      ProcessValue <- "Perfiladores\Perfilador.PL1_1"
   IOField "Champ E/S_115" at 543,307 size 51x25; FormatPattern s999999
      Appearance <- "Perfiladores\Perfilador.PresenciaPieza"
      ProcessValue <- "Perfiladores\Perfilador.PL1_2"
   IOField "Champ E/S_116" at 543,328 size 51x24; FormatPattern s999999
      Appearance <- "Perfiladores\Perfilador.PresenciaPieza"
      ProcessValue <- "Perfiladores\Perfilador.PL2_1"
   IOField "Champ E/S_117" at 543,347 size 51x25; FormatPattern s999999
      Appearance <- "Perfiladores\Perfilador.PresenciaPieza"
      ProcessValue <- "Perfiladores\Perfilador.PL2_2"
   TextField "Campo de texto_123" at 503,310 size 35x18; Text 'PL1-2'
   TextField "Campo de texto_124" at 503,331 size 35x18; Text 'PL2-1'
   TextField "Campo de texto_125" at 503,350 size 35x18; Text 'PL2-2'
   TextField "Campo de texto_134" at 328,210 size 17x18; Text 'F1'
   IOField "Champ E/S_126" at 352,207 size 51x25; FormatPattern s999999
      Appearance <- "Rolos\Rolos.PresenciaPieza"
      ProcessValue <- "Rolos\Rolos.F1"
   IOField "Champ E/S_127" at 352,227 size 51x25; FormatPattern s999999
      Appearance <- "Rolos\Rolos.PresenciaPieza"
      ProcessValue <- "Rolos\Rolos.F2"
   IOField "Champ E/S_128" at 352,248 size 51x24; FormatPattern s999999
      Appearance <- "Rolos\Rolos.PresenciaPieza"
      ProcessValue <- "Rolos\Rolos.F3"
   IOField "Champ E/S_129" at 352,267 size 51x25; FormatPattern s999999
      Appearance <- "Rolos\Rolos.PresenciaPieza"
      ProcessValue <- "Rolos\Rolos.F4"
   TextField "Campo de texto_135" at 328,229 size 17x18; Text 'F2'
   TextField "Campo de texto_136" at 328,249 size 17x18; Text 'F3'
   TextField "Campo de texto_137" at 328,269 size 17x18; Text 'F4'
   TextField "Campo de texto_138" at 328,290 size 35x18; Text 'PL1-1'
   IOField "Champ E/S_130" at 368,287 size 51x25; FormatPattern s999999
      Appearance <- "Rolos\Rolos.PresenciaPieza"
      ProcessValue <- "Rolos\Rolos.PL1_1"
   IOField "Champ E/S_131" at 368,307 size 51x25; FormatPattern s999999
      Appearance <- "Rolos\Rolos.PresenciaPieza"
      ProcessValue <- "Rolos\Rolos.PL1_2"
   IOField "Champ E/S_132" at 368,328 size 51x24; FormatPattern s999999
      Appearance <- "Rolos\Rolos.PresenciaPieza"
      ProcessValue <- "Rolos\Rolos.PL2_1"
   IOField "Champ E/S_133" at 368,347 size 51x25; FormatPattern s999999
      Appearance <- "Rolos\Rolos.PresenciaPieza"
      ProcessValue <- "Rolos\Rolos.PL2_2"
   TextField "Campo de texto_139" at 328,310 size 35x18; Text 'PL1-2'
   TextField "Campo de texto_140" at 328,331 size 35x18; Text 'PL2-1'
   TextField "Campo de texto_141" at 328,350 size 35x18; Text 'PL2-2'
   TextField "Campo de texto_142" at 151,210 size 17x18; Text 'F1'
   IOField "Champ E/S_134" at 175,207 size 51x25; FormatPattern s999999
      Appearance <- "Araña\Araña.PresenciaPieza"
      ProcessValue <- "Araña\Araña.F1"
   IOField "Champ E/S_135" at 175,227 size 51x25; FormatPattern s999999
      Appearance <- "Araña\Araña.PresenciaPieza"
      ProcessValue <- "Araña\Araña.F2"
   IOField "Champ E/S_136" at 175,248 size 51x24; FormatPattern s999999
      Appearance <- "Araña\Araña.PresenciaPieza"
      ProcessValue <- "Araña\Araña.F3"
   IOField "Champ E/S_137" at 175,267 size 51x25; FormatPattern s999999
      Appearance <- "Araña\Araña.PresenciaPieza"
      ProcessValue <- "Araña\Araña.F4"
   TextField "Campo de texto_143" at 151,229 size 17x18; Text 'F2'
   TextField "Campo de texto_144" at 151,249 size 17x18; Text 'F3'
   TextField "Campo de texto_145" at 151,269 size 17x18; Text 'F4'
   TextField "Campo de texto_146" at 151,290 size 35x18; Text 'PL1-1'
   IOField "Champ E/S_138" at 191,287 size 51x25; FormatPattern s999999
      Appearance <- "Araña\Araña.PresenciaPieza"
      ProcessValue <- "Araña\Araña.PL1_1"
   IOField "Champ E/S_139" at 191,307 size 51x25; FormatPattern s999999
      Appearance <- "Araña\Araña.PresenciaPieza"
      ProcessValue <- "Araña\Araña.PL1_2"
   IOField "Champ E/S_140" at 191,328 size 51x24; FormatPattern s999999
      Appearance <- "Araña\Araña.PresenciaPieza"
      ProcessValue <- "Araña\Araña.PL2_1"
   IOField "Champ E/S_141" at 191,347 size 51x25; FormatPattern s999999
      Appearance <- "Araña\Araña.PresenciaPieza"
      ProcessValue <- "Araña\Araña.PL2_2"
   TextField "Campo de texto_147" at 151,310 size 35x18; Text 'PL1-2'
   TextField "Campo de texto_148" at 151,331 size 35x18; Text 'PL2-1'
   TextField "Campo de texto_149" at 151,350 size 35x18; Text 'PL2-2'
   TextField "Campo de texto_150" at 679,210 size 17x18; Text 'F1'
   IOField "Champ E/S_142" at 703,207 size 51x25; FormatPattern s999999
      Appearance <- "Cinta\Cinta.PresenciaPieza"
      ProcessValue <- "Cinta\Cinta.F1"
   IOField "Champ E/S_143" at 703,227 size 51x25; FormatPattern s999999
      Appearance <- "Cinta\Cinta.PresenciaPieza"
      ProcessValue <- "Cinta\Cinta.F2"
   IOField "Champ E/S_144" at 703,248 size 51x24; FormatPattern s999999
      Appearance <- "Cinta\Cinta.PresenciaPieza"
      ProcessValue <- "Cinta\Cinta.F3"
   IOField "Champ E/S_145" at 703,267 size 51x25; FormatPattern s999999
      Appearance <- "Cinta\Cinta.PresenciaPieza"
      ProcessValue <- "Cinta\Cinta.F4"
   TextField "Campo de texto_151" at 679,229 size 17x18; Text 'F2'
   TextField "Campo de texto_152" at 679,249 size 17x18; Text 'F3'
   TextField "Campo de texto_153" at 679,269 size 17x18; Text 'F4'
   TextField "Campo de texto_154" at 679,290 size 35x18; Text 'PL1-1'
   IOField "Champ E/S_146" at 719,287 size 51x25; FormatPattern s999999
      Appearance <- "Cinta\Cinta.PresenciaPieza"
      ProcessValue <- "Cinta\Cinta.PL1_1"
   IOField "Champ E/S_147" at 719,307 size 51x25; FormatPattern s999999
      Appearance <- "Cinta\Cinta.PresenciaPieza"
      ProcessValue <- "Cinta\Cinta.PL1_2"
   IOField "Champ E/S_148" at 719,328 size 51x24; FormatPattern s999999
      Appearance <- "Cinta\Cinta.PresenciaPieza"
      ProcessValue <- "Cinta\Cinta.PL2_1"
   IOField "Champ E/S_149" at 719,347 size 51x25; FormatPattern s999999
      Appearance <- "Cinta\Cinta.PresenciaPieza"
      ProcessValue <- "Cinta\Cinta.PL2_2"
   TextField "Campo de texto_155" at 679,310 size 35x18; Text 'PL1-2'
   TextField "Campo de texto_156" at 679,331 size 35x18; Text 'PL2-1'
   TextField "Campo de texto_157" at 679,350 size 35x18; Text 'PL2-2'
   TextField "Campo de texto_158" at 851,210 size 17x18; Text 'F1'
   IOField "Champ E/S_150" at 875,207 size 51x25; FormatPattern s999999
      Appearance <- "Pinza\Pinza.PresenciaPieza"
      ProcessValue <- "Pinza\Pinza.F1"
   IOField "Champ E/S_151" at 875,227 size 51x25; FormatPattern s999999
      Appearance <- "Pinza\Pinza.PresenciaPieza"
      ProcessValue <- "Pinza\Pinza.F2"
   IOField "Champ E/S_152" at 875,248 size 51x24; FormatPattern s999999
      Appearance <- "Pinza\Pinza.PresenciaPieza"
      ProcessValue <- "Pinza\Pinza.F3"
   IOField "Champ E/S_153" at 875,267 size 51x25; FormatPattern s999999
      Appearance <- "Pinza\Pinza.PresenciaPieza"
      ProcessValue <- "Pinza\Pinza.F4"
   TextField "Campo de texto_159" at 851,229 size 17x18; Text 'F2'
   TextField "Campo de texto_160" at 851,249 size 17x18; Text 'F3'
   TextField "Campo de texto_161" at 851,269 size 17x18; Text 'F4'
   TextField "Campo de texto_162" at 851,290 size 35x18; Text 'PL1-1'
   IOField "Champ E/S_154" at 891,287 size 51x25; FormatPattern s999999
      Appearance <- "Pinza\Pinza.PresenciaPieza"
      ProcessValue <- "Pinza\Pinza.PL1_1"
   IOField "Champ E/S_155" at 891,307 size 51x25; FormatPattern s999999
      Appearance <- "Pinza\Pinza.PresenciaPieza"
      ProcessValue <- "Pinza\Pinza.PL1_2"
   IOField "Champ E/S_156" at 891,328 size 51x24; FormatPattern s999999
      Appearance <- "Pinza\Pinza.PresenciaPieza"
      ProcessValue <- "Pinza\Pinza.PL2_1"
   IOField "Champ E/S_157" at 891,347 size 51x25; FormatPattern s999999
      Appearance <- "Pinza\Pinza.PresenciaPieza"
      ProcessValue <- "Pinza\Pinza.PL2_2"
   TextField "Campo de texto_163" at 851,310 size 35x18; Text 'PL1-2'
   TextField "Campo de texto_164" at 851,331 size 35x18; Text 'PL2-1'
   TextField "Campo de texto_165" at 851,350 size 35x18; Text 'PL2-2'
   TextField "Campo de texto_166" at 1029,210 size 17x18; Text 'F1'
   IOField "Champ E/S_158" at 1053,207 size 51x25; FormatPattern s999999
      Appearance <- "Plegadora\Plegadora.PresenciaPieza"
      ProcessValue <- "Plegadora\Plegadora.F1"
   IOField "Champ E/S_159" at 1053,227 size 51x25; FormatPattern s999999
      Appearance <- "Plegadora\Plegadora.PresenciaPieza"
      ProcessValue <- "Plegadora\Plegadora.F2"
   IOField "Champ E/S_160" at 1053,248 size 51x24; FormatPattern s999999
      Appearance <- "Plegadora\Plegadora.PresenciaPieza"
      ProcessValue <- "Plegadora\Plegadora.F3"
   IOField "Champ E/S_161" at 1053,267 size 51x25; FormatPattern s999999
      Appearance <- "Plegadora\Plegadora.PresenciaPieza"
      ProcessValue <- "Plegadora\Plegadora.F4"
   TextField "Campo de texto_167" at 1029,229 size 17x18; Text 'F2'
   TextField "Campo de texto_168" at 1029,249 size 17x18; Text 'F3'
   TextField "Campo de texto_169" at 1029,269 size 17x18; Text 'F4'
   TextField "Campo de texto_170" at 1029,290 size 35x18; Text 'PL1-1'
   IOField "Champ E/S_162" at 1069,287 size 51x25; FormatPattern s999999
      Appearance <- "Plegadora\Plegadora.PresenciaPieza"
      ProcessValue <- "Plegadora\Plegadora.PL1_1"
   IOField "Champ E/S_163" at 1069,307 size 51x25; FormatPattern s999999
      Appearance <- "Plegadora\Plegadora.PresenciaPieza"
      ProcessValue <- "Plegadora\Plegadora.PL1_2"
   IOField "Champ E/S_164" at 1069,328 size 51x24; FormatPattern s999999
      Appearance <- "Plegadora\Plegadora.PresenciaPieza"
      ProcessValue <- "Plegadora\Plegadora.PL2_1"
   IOField "Champ E/S_165" at 1069,347 size 51x25; FormatPattern s999999
      Appearance <- "Plegadora\Plegadora.PresenciaPieza"
      ProcessValue <- "Plegadora\Plegadora.PL2_2"
   TextField "Campo de texto_171" at 1029,310 size 35x18; Text 'PL1-2'
   TextField "Campo de texto_172" at 1029,331 size 35x18; Text 'PL2-1'
   TextField "Campo de texto_173" at 1029,350 size 35x18; Text 'PL2-2'
   IOField "Champ E/S_32" at 505,100 size 80x25; FormatPattern ????????????????????
      Appearance <- "Perfiladores\Perfilador.PresenciaPieza"
      ProcessValue <- "Perfiladores\Perfilador.Nombre"
   IOField "Champ E/S_33" at 330,100 size 80x25; FormatPattern ????????????????????
      Appearance <- "Rolos\Rolos.PresenciaPieza"
      ProcessValue <- "Rolos\Rolos.Nombre"
   IOField "Champ E/S_34" at 153,100 size 80x25; FormatPattern ????????????????????
      Appearance <- "Araña\Araña.PresenciaPieza"
      ProcessValue <- "Araña\Araña.Nombre"
   IOField "Champ E/S_35" at 681,100 size 80x25; FormatPattern ????????????????????
      Appearance <- "Cinta\Cinta.PresenciaPieza"
      ProcessValue <- "Cinta\Cinta.Nombre"
   IOField "Champ E/S_41" at 853,100 size 80x25; FormatPattern ????????????????????
      Appearance <- "Pinza\Pinza.PresenciaPieza"
      ProcessValue <- "Pinza\Pinza.Nombre"
   IOField "Champ E/S_42" at 1031,100 size 80x25; FormatPattern ????????????????????
      Appearance <- "Plegadora\Plegadora.PresenciaPieza"
      ProcessValue <- "Plegadora\Plegadora.Nombre"
   TextField "Campo de texto_67" at 143,608 size 33x18; Text 'E2H2'
   IOField "Champ E/S_29" at 221,605 size 85x25; FormatPattern s9999999999
      ProcessValue <- "Pos_E2H2"
      Appearance <- "Pinza\Pinza.PresenciaPieza"
   IOField "Champ E/S_30" at 221,625 size 85x25; FormatPattern s9999999999
      ProcessValue <- "Pos_Entrega"
      Appearance <- "Pinza\Pinza.PresenciaPieza"
   TextField "Campo de texto_68" at 143,627 size 47x18; Text 'Entrega'
   IOField "Champ E/S_31" at 305,605 size 85x25; FormatPattern s9999999999
      ProcessValue <- "Pos_E2H2(3)"
      Appearance <- "Pinza\Pinza.PresenciaPieza"
   IOField "Champ E/S_36" at 305,625 size 85x25; FormatPattern s9999999999
      ProcessValue <- "Pos_Entrega(3)"
      Appearance <- "Pinza\Pinza.PresenciaPieza"
   IOField "Champ E/S_61" at 608,605 size 85x25; FormatPattern s9999999999
      ProcessValue <- "Pos_E2H2(1)"
      Appearance <- "Pinza\Pinza.PresenciaPieza"
   IOField "Champ E/S_62" at 608,625 size 85x25; FormatPattern s9999999999
      ProcessValue <- "Pos_Entrega(1)"
      Appearance <- "Pinza\Pinza.PresenciaPieza"
   IOField "Champ E/S_73" at 690,605 size 85x25; FormatPattern s9999999999
      ProcessValue <- "Pos_E2H2(4)"
      Appearance <- "Pinza\Pinza.PresenciaPieza"
   IOField "Champ E/S_74" at 690,625 size 85x25; FormatPattern s9999999999
      ProcessValue <- "Pos_Entrega(4)"
      Appearance <- "Pinza\Pinza.PresenciaPieza"
   IOField "Champ E/S_85" at 995,605 size 85x25; FormatPattern s9999999999
      ProcessValue <- "Pos_E2H2(2)"
      Appearance <- "Pinza\Pinza.PresenciaPieza"
   IOField "Champ E/S_86" at 995,625 size 85x25; FormatPattern s9999999999
      ProcessValue <- "Pos_Entrega(2)"
      Appearance <- "Pinza\Pinza.PresenciaPieza"
   IOField "Champ E/S_97" at 1077,605 size 85x25; FormatPattern s9999999999
      ProcessValue <- "Pos_E2H2(5)"
      Appearance <- "Pinza\Pinza.PresenciaPieza"
   IOField "Champ E/S_98" at 1077,625 size 85x25; FormatPattern s9999999999
      ProcessValue <- "Pos_Entrega(5)"
      Appearance <- "Pinza\Pinza.PresenciaPieza"
   TextField "Campo de texto_69" at 534,608 size 33x18; Text 'E2H2'
   TextField "Campo de texto_70" at 534,627 size 47x18; Text 'Entrega'
   TextField "Campo de texto_71" at 917,608 size 33x18; Text 'E2H2'
   TextField "Campo de texto_72" at 917,627 size 47x18; Text 'Entrega'

Template "Template" 1280x770
   TextField "Template_Plantilla_Campo de texto" at 0,0 size 1280x24; Text 'Movimiento Manual Seleccionado -'
      Visibility <- "DB_OP.RC1"
   TextField "Template_Plantilla_Campo de texto_0" at 0,-1 size 1280x24; Text 'Movimiento Manual Seleccionado -'
      Visibility <- "DB_OP.RC2"
   Button "Template_Plantilla_Bouton_1" at 278,715 size 150x53; TextOff 'SEGUIMIENTO DE DATOS SYSTEM'
      on Click: ActivateScreen("eProC - Seguimiento Datos", 0)
   Button "Template_Plantilla_Bouton_0" at 1085,715 size 193x53; TextOff 'ALARMAS / DEFAUT'
      on Press: ActivateScreen("eProC - Alarmas", 0)
   Button "Template_Plantilla_Botón_2" at 573,715 size 70x53; TextOff 'Text'; Authorization "Nivel 2"; PictureOn "Usuario"; PictureOff "Usuario"
      on Activate: ActivateScreen("Gesión de Usuarios", 0)
   Button "Template_Plantilla_Botón_3" at 129,715 size 150x53; TextOff 'SELECCIÓN RECETAS'
      on Click: ActivateScreen("eProC - Recetas", 0)
   Button "Template_Plantilla_Botón_4" at 641,715 size 150x53; TextOff 'Text'
   SymbolicIOField "Template_Plantilla_Campo ES simbólico" at 234,0 size 896x24; TextOff '0'; TextOn '1'; TextList "RC2"
      ProcessValue <- "DB_OP.RC2"
      Visibility <- "DB_OP.RC2"
   SymbolicIOField "Template_Plantilla_Campo ES simbólico_0" at 234,0 size 896x24; TextOff '0'; TextOn '1'; TextList "RC1"
      ProcessValue <- "DB_OP.RC1"
      Visibility <- "DB_OP.RC1"
   Button "Plantilla_Botón_1" at 1,715 size 130x53; TextOff 'PRINCIPAL'
      on Click: ActivateScreen("eProC - Principal", 0)
   SymbolicIOField "Template_Plantilla_Campo ES simbólico_1" at 0,0 size 1280x24; TextOff '0'; TextOn '1'; TextList "Warnings"
      ProcessValue <- "Warnings"
      Visibility <- "Warning Activo"
   Button "Template_Plantilla_Botón_5" at 789,715 size 150x53; TextOff 'Text'
   Button "Template_Plantilla_Botón_6" at 937,715 size 150x53; TextOff 'Text'
   Button "Template_Plantilla_Bouton_2" at 1085,715 size 193x53; TextOff 'ALARMAS / DEFAUT'
      on Press: ActivateScreen("eProC - Alarmas", 0)
      Visibility <- "DB_OP.P_DEFAUT"
   Button "Template_Plantilla_Botón_1" at 424,715 size 150x53; TextOff 'Text'

PopupScreen "Configurador de Recetas" 1010x320
   Rectangle "Rectángulo_15" at 0,0 size 1010x320
      Visibility <- "Receta\VerHeladera"
   TextField "Campo de texto_55" at 26,93 size 17x26; Text 'A'
      Visibility <- "Receta\VerHeladera"
   IOField "Champ E/S_42" at 40,95 size 88x23; FormatPattern 9999999
      ProcessValue <- "Receta\Recetas.A"
      Visibility <- "Receta\VerHeladera"
   IOField "Champ E/S_43" at 219,31 size 74x23; FormatPattern 9999999
      ProcessValue <- "Receta\Recetas.B"
      Visibility <- "Receta\VerHeladera"
   IOField "Champ E/S_44" at 115,31 size 74x23; FormatPattern 9999999
      Visibility <- "Receta\VerHeladera"
      ProcessValue <- "Receta\Recetas.C"
   IOField "Champ E/S_45" at 40,229 size 88x24; FormatPattern 9999999
      ProcessValue <- "Receta\Recetas.D"
      Visibility <- "Receta\VerHeladera"
   IOField "Champ E/S_46" at 56,138 size 72x24; FormatPattern 99999
      ProcessValue <- "Receta\Recetas.F2"
      Visibility <- "Receta\VerHeladera"
   IOField "Champ E/S_47" at 54,273 size 74x23; FormatPattern 99999
      ProcessValue <- "Receta\Recetas.F1"
      Visibility <- "Receta\VerHeladera"
   IOField "Champ E/S_48" at 331,273 size 70x23; FormatPattern 99999
      ProcessValue <- "Receta\Recetas.F3"
      Visibility <- "Receta\VerHeladera"
   IOField "Champ E/S_49" at 56,117 size 72x24; FormatPattern 99999
      Visibility <- "Receta\VerHeladera"
      ProcessValue <- "Receta\OFFSET.RECETTE.OFFSET_PL1_1"
   IOField "Champ E/S_50" at 58,250 size 75x24; FormatPattern 99999
      Visibility <- "Receta\VerHeladera"
      ProcessValue <- "Receta\OFFSET.RECETTE.OFFSET_PL1_2"
   IOField "Champ E/S_51" at 355,251 size 70x24; FormatPattern 99999
      ProcessValue <- "Receta\Recetas.PL2_1"
      Visibility <- "Receta\VerHeladera"
   TextField "Campo de texto_56" at 202,29 size 17x26; Text 'B'
      Visibility <- "Receta\VerHeladera"
   TextField "Campo de texto_57" at 98,29 size 17x26; Text 'C'
      Visibility <- "Receta\VerHeladera"
   TextField "Campo de texto_58" at 27,226 size 19x26; Text 'D'
      Visibility <- "Receta\VerHeladera"
   Polygon "Polígono_12" at 165,79 size 110x27
      Visibility <- "Receta\VerHeladera"
   Polygon "Polígono_13" at 168,106 size 42x119
      Visibility <- "Receta\VerHeladera"
   Polygon "Polígono_14" at 163,207 size 66x19
      Visibility <- "Receta\VerHeladera"
   Polyline "Línea poligonal_2" at 123,226 size 42x13
      Visibility <- "Receta\VerHeladera"
   Polyline "Línea poligonal_3" at 123,109 size 38x0
      Visibility <- "Receta\VerHeladera"
   IOField "Champ E/S_52" at 328,229 size 88x24; FormatPattern 9999999
      ProcessValue <- "Receta\Recetas.D"
      Visibility <- "Receta\VerHeladera"
   TextField "Campo de texto_60" at 310,226 size 19x26; Text 'D'
      Visibility <- "Receta\VerHeladera"
   Polyline "Línea poligonal_10" at 234,227 size 64x12
      Visibility <- "Receta\VerHeladera"
   Polyline "Línea poligonal_4" at 149,55 size 40x36
      Visibility <- "Receta\VerHeladera"
   Polyline "Línea poligonal_5" at 238,53 size 0x25
      Visibility <- "Receta\VerHeladera"
   Polygon "Polígono_15" at 211,207 size 66x19
      Visibility <- "Receta\VerHeladera"
   Polygon "Polígono_16" at 234,79 size 43x145
      Visibility <- "Receta\VerHeladera"
   IOField "Champ E/S_53" at 330,137 size 70x25; FormatPattern 99999
      ProcessValue <- "Receta\Recetas.F4"
      Visibility <- "Receta\VerHeladera"
   IOField "Champ E/S_54" at 352,117 size 69x24; FormatPattern 99999
      ProcessValue <- "Receta\Recetas.PL2_2"
      Visibility <- "Receta\VerHeladera"
   TextField "Campo de texto_62" at 306,93 size 17x26; Text 'A'
      Visibility <- "Receta\VerHeladera"
   IOField "Champ E/S_55" at 325,95 size 86x23; FormatPattern 9999999
      ProcessValue <- "Receta\Recetas.A"
      Visibility <- "Receta\VerHeladera"
   Polyline "Línea poligonal_7" at 238,109 size 59x0
      Visibility <- "Receta\VerHeladera"
   TextField "Campo de texto_63" at 13,117 size 40x22; Text 'PL1-2'
      Visibility <- "Receta\VerHeladera"
   TextField "Campo de texto_64" at 38,138 size 20x22; Text 'F2'
      Visibility <- "Receta\VerHeladera"
   TextField "Campo de texto_65" at 14,250 size 40x22; Text 'PL1-1'
      Visibility <- "Receta\VerHeladera"
   TextField "Campo de texto_66" at 38,273 size 20x22; Text 'F1'
      Visibility <- "Receta\VerHeladera"
   TextField "Campo de texto_67" at 306,117 size 40x22; Text 'PL2-2'
      Visibility <- "Receta\VerHeladera"
   TextField "Campo de texto_68" at 309,138 size 20x22; Text 'F4'
      Visibility <- "Receta\VerHeladera"
   TextField "Campo de texto_69" at 309,251 size 40x22; Text 'PL2-1'
      Visibility <- "Receta\VerHeladera"
   TextField "Campo de texto_70" at 310,273 size 20x22; Text 'F3'
      Visibility <- "Receta\VerHeladera"
   RecipeView "RecipeView" at 456,70 size 539x71; RecipeNameCaption 'Receta:'; DataRecordNameCaption 'Receta:'; ValueCaption 'Valor'; RecipeNrCaption 'N.º:'; DataRecordNrCaption 'Nº:'; EntryNameCaption 'Nombre de entrada'; Tag4DataRecord "Receta\Recetas.Nombre"; Recipe "Pieza"
      Visibility <- "Receta\VerHeladera"
   Button "Botón_7" at 891,17 size 90x43; TextOff 'Cerrar'
      on Click: InvertBit("Receta\VerHeladera"); ResetBit("Receta Almacén1\VerHeladera"); ResetBit("Receta Almacén 2\VerHeladera"); ResetBit("Receta Almacén1\Detalles"); ResetBit("Receta Almacén 2\Detalles"); function_efd93a16("Configurador de Recetas", 0, 0, -1, -1, 1)
      Visibility <- "Receta\VerHeladera"
   Rectangle "Rectángulo_12" at 474,210 size 502x92
      Visibility <- "Receta\VerHeladera"
   Polygon "Polígono_2" at 792,262 size 22x25
      Visibility <- "Receta Almacén1\CA_KM01_1"
   IOField "Champ E/S_28" at 898,261 size 64x32; FormatPattern 9999
      ProcessValue <- "DB_OP.M1_P_CPT"
   IOField "Champ E/S_29" at 898,222 size 64x32; FormatPattern 9999
      ProcessValue <- "DB_OP.M2_P_CPT"
   IOField "Champ E/S_30" at 822,261 size 61x32; FormatPattern 9999
      ProcessValue <- "DB_OP.M1_V_CPT"
   IOField "Champ E/S_31" at 822,222 size 61x32; FormatPattern 9999
      ProcessValue <- "DB_OP.M2_V_CPT"
   Polygon "Polígono_4" at 792,225 size 21x24
      Visibility <- "Receta Almacén 2\CA_KM01_2"
   Button "Button_6" at 490,258 size 82x35; TextOff 'Cargar'; PictureOff "Flèche_Droite"
      on Press: function_eba64363('REFERENCE', "Receta\Recetas.Nombre", 1, N)
      on Release: SetBit("Receta\Recetas.x_M1")
      Visibility <- "Receta\VerHeladera"
      Appearance <- "Receta\Recetas.x_M1"
   Button "Button_7" at 490,221 size 82x33; TextOff 'Cargar'; PictureOff "Flèche_Droite"
      on Press: function_eba64363('REFERENCE', "Receta\Recetas.Nombre", 1, N)
      on Release: SetBit("Receta\Recetas.x_M2")
      Visibility <- "Receta\VerHeladera"
      Appearance <- "Receta\Recetas.x_M2"
   TextField "Campo de texto_14" at 587,265 size 72x22; Text 'Almacén 1'
   IOField "Champ E/S_56" at 675,265 size 120x24; FormatPattern ??????????
      ProcessValue <- "Receta Almacén1\Recetas.REC_MG1.NOM"
   TextField "Campo de texto_15" at 587,226 size 72x22; Text 'Almacén 2'
   IOField "Champ E/S_57" at 675,226 size 118x24; FormatPattern ??????????
      ProcessValue <- "Receta Almacén 2\Recetas.REC_MG2.NOM"
   TextField "Campo de texto_59" at 470,50 size 164x26; Text 'Selección de Modelo'
      Visibility <- "Receta\VerHeladera"

PopupScreen "Comandos Araña" 1280x714
   Circle "Cercle_11" at 358,354 size 13x13
      Appearance <- "25S8"
   Circle "Cercle_12" at 359,303 size 13x13
      Appearance <- "25S7"
   Circle "Cercle_0" at 358,375 size 13x13
      Appearance <- "25S4"
   Circle "Cercle_1" at 398,262 size 12x12
      Appearance <- "25S3"
   Circle "Cercle_2" at 320,381 size 12x12
      Appearance <- "25S5"
   Circle "Cercle_3" at 399,300 size 12x12
      Appearance <- "26S3"
   TextField "Campo de texto_1" at 509,184 size 154x18; Text '25S3 - Fin de Carrera Arriba'
   TextField "Campo de texto_6" at 94,362 size 154x18; Text '25S5 - Fin de Carrera Abajo'
   TextField "Campo de texto_10" at 515,231 size 176x18; Text '26S3 - En Posición de Descarga'
   TextField "Campo de texto_8" at 105,226 size 148x18; Text '25S7 - Pistón 2 Expandido'
   TextField "Campo de texto_18" at 107,270 size 144x18; Text '25S8 - Pistón 2 Contraído'
   TextField "Campo de texto_19" at 107,326 size 144x18; Text '25S4 - Pistón 1 Contraído'
   TextField "Campo de texto_20" at 521,268 size 110x18; Text '25S6 - Araña Abajo'
   Circle "Cercle_5" at 401,347 size 13x13
      Appearance <- "25S6"
   Circle "Cercle" at 340,467 size 13x13
      Appearance <- "26S1"
   TextField "Campo de texto_9" at 91,496 size 204x18; Text '26S1 - Tulipas Apoyadas en la Chapa'
   TextField "Campo de texto_21" at 657,356 size 126x18; Text '26S5 - Bajar Velocidad'
   TextField "Campo de texto_22" at 652,316 size 176x18; Text '26S3 - En Posición de Descarga'
   TextField "Campo de texto_23" at 653,421 size 170x46; Text 'M03 - Motor Transporte Araña KM02.1 -> Hacia Rolos KM02.2 -> Hacia Almacenes'
   TextField "Campo de texto_24" at 672,505 size 126x18; Text '26S4 - Bajar Velocidad'
   TextField "Campo de texto_25" at 678,546 size 157x18; Text '26S2 - En Posición de Carga'
   Circle "Cercle_4" at 572,534 size 12x12
      Appearance <- "26S2"
   Circle "Cercle_6" at 567,494 size 12x12
      Appearance <- "26S4"
   Circle "Cercle_7" at 554,342 size 12x12
      Appearance <- "26S5"
   Circle "Cercle_8" at 549,303 size 12x12
      Appearance <- "26S3"
   Polygon "Polígono_3" at 206,439 size 325x50
      Visibility <- "Araña\Araña.PresenciaPieza"
   Rectangle "Rectángulo_7" at 989,250 size 248x208
      Visibility <- "MANU"
   Rectangle "Rectángulo_12" at 989,246 size 248x29
      Visibility <- "MANU"
   Rectangle "Rectángulo_9" at 843,27 size 118x128
      Visibility <- "MANU"
   Rectangle "Rectángulo_8" at 843,27 size 118x29
      Visibility <- "MANU"
   TextField "Campo de texto_3" at 870,31 size 64x18; Text 'Transporte'
      Visibility <- "MANU"
   TextField "Campo de texto_11" at 1010,252 size 66x18; Text 'Aire Tulipas'
      Visibility <- "MANU"
   Button "Botón_4" at 859,71 size 88x33; TextOff 'Avance'
      on Press: SetTag("DB_OP.RC1", 11); SetBit("DB_OP.OP_SELMANU1")
      Visibility <- "MANU"
      Appearance <- "DB_OP.RC1"
   Button "Botón_5" at 859,109 size 88x33; TextOff 'Retroceso'
      on Press: SetTag("DB_OP.RC1", 12); SetBit("DB_OP.OP_SELMANU1")
      Visibility <- "MANU"
      Appearance <- "DB_OP.RC1"
   Button "Botón_10" at 1065,290 size 72x33; TextOff 'Activar'
      on Press: SetTag("DB_OP.RC1", 20); SetBit("DB_OP.OP_SELMANU1")
      Visibility <- "MANU"
      Appearance <- "DB_OP.RC1"
   Button "Botón_17" at 1145,290 size 72x33; TextOff 'Desactivar'
      on Press: SetTag("DB_OP.RC1", 21); SetBit("DB_OP.OP_SELMANU1")
      Visibility <- "MANU"
      Appearance <- "DB_OP.RC1"
   TextField "Campo de texto_12" at 1010,296 size 37x18; Text 'Todas'
      Visibility <- "MANU"
   Button "Botón_1" at 1065,336 size 72x33; TextOff 'Activar'
      on Press: SetTag("DB_OP.RC1", 32); SetBit("DB_OP.OP_SELMANU1")
      Visibility <- "MANU"
      Appearance <- "DB_OP.RC1"
   Button "Botón_23" at 1065,373 size 72x33; TextOff 'Activar'
      on Press: SetTag("DB_OP.RC1", 34); SetBit("DB_OP.OP_SELMANU1")
      Visibility <- "MANU"
      Appearance <- "DB_OP.RC1"
   Button "Botón_24" at 1065,411 size 72x33; TextOff 'Activar'
      on Press: SetTag("DB_OP.RC1", 36); SetBit("DB_OP.OP_SELMANU1")
      Visibility <- "MANU"
      Appearance <- "DB_OP.RC1"
   Button "Botón_26" at 1145,336 size 72x33; TextOff 'Desactivar'
      on Press: SetTag("DB_OP.RC1", 33); SetBit("DB_OP.OP_SELMANU1")
      Visibility <- "MANU"
      Appearance <- "DB_OP.RC1"
   Button "Botón_27" at 1145,373 size 72x33; TextOff 'Desactivar'
      on Press: SetTag("DB_OP.RC1", 35); SetBit("DB_OP.OP_SELMANU1")
      Visibility <- "MANU"
      Appearance <- "DB_OP.RC1"
   Button "Botón_28" at 1145,411 size 72x33; TextOff 'Desactivar'
      on Press: SetTag("DB_OP.RC1", 37); SetBit("DB_OP.OP_SELMANU1")
      Visibility <- "MANU"
      Appearance <- "DB_OP.RC1"
   TextField "Campo de texto_2" at 1008,343 size 48x18; Text 'Grupo 1'
      Visibility <- "MANU"
   TextField "Campo de texto_4" at 1008,381 size 48x18; Text 'Grupo 2'
      Visibility <- "MANU"
   TextField "Campo de texto_5" at 1008,419 size 48x18; Text 'Grupo 3'
      Visibility <- "MANU"
   Rectangle "Rectángulo_1" at 989,483 size 248x208
      Visibility <- "MANU"
   Rectangle "Rectángulo_2" at 989,479 size 248x29
      Visibility <- "MANU"
   TextField "Campo de texto_13" at 1010,485 size 74x18; Text 'Vacío Tulipas'
      Visibility <- "MANU"
   TextField "Campo de texto_14" at 1010,529 size 37x18; Text 'Todas'
      Visibility <- "MANU"
   TextField "Campo de texto_15" at 1008,576 size 48x18; Text 'Grupo 1'
      Visibility <- "MANU"
   TextField "Campo de texto_16" at 1008,614 size 48x18; Text 'Grupo 2'
      Visibility <- "MANU"
   TextField "Campo de texto_17" at 1008,652 size 48x18; Text 'Grupo 3'
      Visibility <- "MANU"
   Button "Botón_21" at 1065,523 size 72x33; TextOff 'Activar'
      on Press: SetTag("DB_OP.RC1", 30); SetBit("DB_OP.OP_SELMANU1")
      Visibility <- "MANU"
      Appearance <- "DB_OP.RC1"
   Button "Botón_25" at 1145,523 size 72x33; TextOff 'Desactivar'
      on Press: SetTag("DB_OP.RC1", 31); SetBit("DB_OP.OP_SELMANU1")
      Visibility <- "MANU"
      Appearance <- "DB_OP.RC1"
   Button "Botón_14" at 1065,569 size 72x33; TextOff 'Activar'
      on Press: SetTag("DB_OP.RC1", 22); SetBit("DB_OP.OP_SELMANU1")
      Visibility <- "MANU"
      Appearance <- "DB_OP.RC1"
   Button "Botón_15" at 1065,606 size 72x33; TextOff 'Activar'
      on Press: SetTag("DB_OP.RC1", 24); SetBit("DB_OP.OP_SELMANU1")
      Visibility <- "MANU"
      Appearance <- "DB_OP.RC1"
   Button "Botón_16" at 1065,644 size 72x33; TextOff 'Activar'
      on Press: SetTag("DB_OP.RC1", 26); SetBit("DB_OP.OP_SELMANU1")
      Visibility <- "MANU"
      Appearance <- "DB_OP.RC1"
   Button "Botón_18" at 1145,569 size 72x33; TextOff 'Desactivar'
      on Press: SetTag("DB_OP.RC1", 23); SetBit("DB_OP.OP_SELMANU1")
      Visibility <- "MANU"
      Appearance <- "DB_OP.RC1"
   Button "Botón_19" at 1145,606 size 72x33; TextOff 'Desactivar'
      on Press: SetTag("DB_OP.RC1", 25); SetBit("DB_OP.OP_SELMANU1")
      Visibility <- "MANU"
      Appearance <- "DB_OP.RC1"
   Button "Botón_20" at 1145,644 size 72x33; TextOff 'Desactivar'
      on Press: SetTag("DB_OP.RC1", 27); SetBit("DB_OP.OP_SELMANU1")
      Visibility <- "MANU"
      Appearance <- "DB_OP.RC1"
   Rectangle "Rectángulo_10" at 988,26 size 248x201
      Visibility <- "MANU"
   Button "Botón_6" at 1012,65 size 202x33; TextOff 'Subir (Pistón Superior)'
      on Press: SetTag("DB_OP.RC1", 16); SetBit("DB_OP.OP_SELMANU1")
      Visibility <- "MANU"
      Appearance <- "DB_OP.RC1"
   Button "Botón_7" at 1012,103 size 202x33; TextOff 'Bajar (Pistón Superior)'
      on Press: SetTag("DB_OP.RC1", 15); SetBit("DB_OP.OP_SELMANU1")
      Visibility <- "MANU"
      Appearance <- "DB_OP.RC1"
   Button "Botón_8" at 1012,179 size 202x33; TextOff 'Bajar (Pistón Inferior)'
      on Press: SetTag("DB_OP.RC1", 13); SetBit("DB_OP.OP_SELMANU1")
      Visibility <- "MANU"
      Appearance <- "DB_OP.RC1"
   Button "Botón_9" at 1012,141 size 202x33; TextOff 'Subir (Pistón Inferior)'
      on Press: SetTag("DB_OP.RC1", 14); SetBit("DB_OP.OP_SELMANU1")
      Visibility <- "MANU"
      Appearance <- "DB_OP.RC1"
   Rectangle "Rectángulo_11" at 988,26 size 248x29
      Visibility <- "MANU"
   TextField "Campo de texto_7" at 1056,30 size 110x18; Text 'Movimiento Vertical'
      Visibility <- "MANU"
   GraphicIOField "Campo ES gráfico_1" at 159,226 size 460x334; PictureList "Araña"
      ProcessValue <- "Alarma_Araña"

PopupScreen "Comandos Almacenes" 1280x714
   Rectangle "Rectángulo_9" at 844,194 size 118x128
      Visibility <- "MANU"
   Rectangle "Rectángulo_8" at 844,194 size 118x29
      Visibility <- "MANU"
   TextField "Campo de texto_3" at 860,198 size 86x18; Text 'Intercambiador'
      Visibility <- "MANU"
   Button "Botón_1" at 859,238 size 88x33; TextOff 'Avance'
      on Press: SetTag("DB_OP.RC1", 1); SetBit("DB_OP.OP_SELMANU1")
      Visibility <- "MANU"
      Appearance <- "DB_OP.RC1"
   Button "Botón_2" at 859,276 size 88x33; TextOff 'Retroceso'
      on Press: SetTag("DB_OP.RC1", 2); SetBit("DB_OP.OP_SELMANU1")
      Visibility <- "MANU"
      Appearance <- "DB_OP.RC1"
   Circle "Cercle_1" at 407,425 size 14x14
      Appearance <- "26S6"
   TextField "Campo de texto_2" at 87,557 size 259x22; Text '26S7 - Almacén 2 en puesto de Espera'
   TextField "Campo de texto_4" at 36,478 size 266x22; Text '26S6 - Almacén 2 en puesto de Trabajo'
   GraphicIOField "Campo ES gráfico_2" at 416,233 size 388x286; PictureList "Grupo 1 - Almacén A"
      ProcessValue <- "26S7"
   GraphicIOField "Campo ES gráfico_1" at 416,233 size 388x286; PictureList "Grupo 1 - Almacén B"
      ProcessValue <- "26S7"
      Visibility <- "Alarma_Almacenes"
   Circle "Cercle_2" at 502,466 size 14x14
      Appearance <- "26S7"
   TextField "Campo de texto_6" at 52,590 size 285x22; Text 'M01 - Motor Intercambiador de Almacenes'

PopupScreen "Comandos Rolos" 1280x714
   GraphicIOField "Campo ES gráfico_4" at 134,166 size 538x272; PictureList "Rolos"
      ProcessValue <- "Alarma_Perfiladores"
   Polygon "Polígono_3" at 184,215 size 385x136
      Visibility <- "Rolos\Rolos.PresenciaPieza"
   Rectangle "Rectángulo_9" at 811,197 size 118x128
      Visibility <- "MANU"
   Rectangle "Rectángulo_8" at 811,197 size 118x29
      Visibility <- "MANU"
   TextField "Campo de texto_3" at 854,201 size 32x18; Text 'Rolos'
      Visibility <- "MANU"
   Button "Botón_29" at 826,241 size 88x33; TextOff 'Avance'
      on Press: SetTag("DB_OP.RC1", 41); SetBit("DB_OP.OP_SELMANU1")
      Visibility <- "MANU"
      Appearance <- "DB_OP.RC1"
   Button "Botón_30" at 826,279 size 88x33; TextOff 'Retroceso'
      on Press: SetTag("DB_OP.RC1", 42); SetBit("DB_OP.OP_SELMANU1")
      Visibility <- "MANU"
      Appearance <- "DB_OP.RC1"
   TextField "Campo de texto_7" at 303,476 size 104x32; Text '27S3 - Chapa en Entrada Perfilador'
   Circle "Cercle_10" at 201,328 size 12x12
      Appearance <- "27S3"
   Circle "Cercle_13" at 349,283 size 12x12
      Appearance <- "26S8"
   TextField "Campo de texto_11" at 455,437 size 114x32; Text '26S8 - Chapa en Transporte de Rolos'

PopupScreen "Comandos Piqueteador" 1280x714
   Button "Botón_32" at 397,449 size 118x33; TextOff 'Bajar Tope'
      on Press: SetTag("DB_OP.RC2", 36); SetBit("DB_OP.OP_SELMANU2")
      Visibility <- "MANU"
      Appearance <- "DB_OP.RC2"
   Button "Botón_33" at 397,411 size 118x33; TextOff 'Subir Tope'
      on Press: SetTag("DB_OP.RC2", 35); SetBit("DB_OP.OP_SELMANU2")
      Visibility <- "MANU"
      Appearance <- "DB_OP.RC2"
   Button "Botón_34" at 517,449 size 104x33; TextOff 'Bajar Herr.'
      on Press: SetTag("DB_OP.RC2", 40); SetBit("DB_OP.OP_SELMANU2")
      Visibility <- "MANU"
      Appearance <- "DB_OP.RC2"
   Button "Botón_35" at 517,411 size 104x33; TextOff 'Subir Herr.'
      on Press: SetTag("DB_OP.RC2", 41); SetBit("DB_OP.OP_SELMANU2")
      Visibility <- "MANU"
      Appearance <- "DB_OP.RC2"
   TextField "Campo de texto_5" at 1020,369 size 81x18; Text 'Herramienta 2'
   TextField "Campo de texto_2" at 748,373 size 81x18; Text 'Herramienta 1'
   Button "Botón_20" at 674,411 size 88x33; TextOff 'ON'
      on Press: SetTag("DB_OP.RC2", 42); SetBit("DB_OP.OP_SELMANU2")
      Visibility <- "MANU"
      Appearance <- "DB_OP.RC2"
   Button "Botón_21" at 946,411 size 88x33; TextOff 'ON'
      on Press: SetTag("DB_OP.RC2", 46); SetBit("DB_OP.OP_SELMANU2")
      Visibility <- "MANU"
      Appearance <- "DB_OP.RC2"
   Button "Botón_22" at 764,411 size 88x33; TextOff 'OFF'
      on Press: SetTag("DB_OP.RC2", 43); SetBit("DB_OP.OP_SELMANU2")
      Visibility <- "MANU"
      Appearance <- "DB_OP.RC2"
   Button "Botón_23" at 1036,411 size 88x33; TextOff 'OFF'
      on Press: SetTag("DB_OP.RC2", 47); SetBit("DB_OP.OP_SELMANU2")
      Visibility <- "MANU"
      Appearance <- "DB_OP.RC2"
   Button "Botón_28" at 674,449 size 88x33; TextOff 'ON'
      on Press: SetTag("DB_OP.RC2", 44); SetBit("DB_OP.OP_SELMANU2")
      Visibility <- "MANU"
      Appearance <- "DB_OP.RC2"
   Button "Botón_1" at 946,447 size 88x33; TextOff 'ON'
      on Press: SetTag("DB_OP.RC2", 48); SetBit("DB_OP.OP_SELMANU2")
      Visibility <- "MANU"
      Appearance <- "DB_OP.RC2"
   Button "Botón_2" at 764,449 size 88x33; TextOff 'OFF'
      on Press: SetTag("DB_OP.RC2", 45); SetBit("DB_OP.OP_SELMANU2")
      Visibility <- "MANU"
      Appearance <- "DB_OP.RC2"
   Button "Botón_31" at 1036,447 size 88x33; TextOff 'OFF'
      on Press: SetTag("DB_OP.RC2", 49); SetBit("DB_OP.OP_SELMANU2")
      Visibility <- "MANU"
      Appearance <- "DB_OP.RC2"
   GraphicIOField "Campo ES gráfico_8" at 250,43 size 289x268; PictureList "Formador"
      ProcessValue <- "Alarma_Formador"
   Rectangle "Rectángulo_9" at 930,366 size 254x128
      Visibility <- "MANU"
   Circle "Cercle_6" at 349,49 size 10x10
      Appearance <- "28S5"
   Circle "Cercle_7" at 349,78 size 10x10
      Appearance <- "28S6"
   TextField "Campo de texto_4" at 72,33 size 180x18; Text '28S5 - Herramientas Bloqueadas'
   TextField "Campo de texto_9" at 54,61 size 200x18; Text '28S6 - Herramientas Desbloqueadas'
   Circle "Cercle_8" at 451,121 size 10x10
      Appearance <- "28S3"
   Circle "Cercle_9" at 465,130 size 10x10
      Appearance <- "28S4"
   Circle "Cercle_10" at 518,168 size 10x10
      Appearance <- "28S1"
   Circle "Cercle_16" at 495,149 size 10x10
      Appearance <- "28S2"
   Circle "Cercle_0" at 433,216 size 10x10
      Appearance <- "27S5"
   Circle "Cercle_17" at 410,198 size 10x10
      Appearance <- "27S6"
   Circle "Cercle_18" at 361,163 size 10x10
      Appearance <- "27S7"
   Circle "Cercle_19" at 379,176 size 10x10
      Appearance <- "27S8"
   TextField "Campo de texto_14" at 530,72 size 146x18; Text '28S3 - Herr. 2 Matriz OFF'
   TextField "Campo de texto_15" at 543,91 size 142x18; Text '28S4 - Herr. 2 Matriz ON'
   TextField "Campo de texto_16" at 589,139 size 152x18; Text '28S1 - Herr. 2 Martillo OFF'
   TextField "Campo de texto_17" at 562,118 size 148x18; Text '28S2 - Herr. 2 Martillo ON'
   TextField "Campo de texto_18" at 40,196 size 146x18; Text '27S7 - Herr. 1 Matriz OFF'
   TextField "Campo de texto_19" at 64,219 size 142x18; Text '27S8 - Herr. 1 Matriz ON'
   TextField "Campo de texto_20" at 90,276 size 152x18; Text '27S5 - Herr. 1 Martillo OFF'
   TextField "Campo de texto_21" at 73,257 size 148x18; Text '27S6 - Herr. 1 Martillo ON'
   Rectangle "Rectángulo_1" at 381,369 size 254x128
      Visibility <- "MANU"
   Rectangle "Rectángulo_2" at 381,369 size 254x29
      Visibility <- "MANU"
   TextField "Campo de texto_1" at 491,373 size 45x18; Text 'General'
      Visibility <- "MANU"
   Rectangle "Rectángulo_3" at 658,369 size 254x128
      Visibility <- "MANU"
   IOField "Campo ES_1" at 480,552 size 96x32; FormatPattern 99999999
      ProcessValue <- "PosiciónFormado1"
   IOField "Campo ES_2" at 707,585 size 96x32; FormatPattern 99999999
      ProcessValue <- "PosiciónFormado2"
   IOField "Campo ES_3" at 480,585 size 96x32; FormatPattern 99999999
      ProcessValue <- "PosiciónFormado3"
   IOField "Campo ES_4" at 707,552 size 96x32; FormatPattern 99999999
      ProcessValue <- "PosiciónFormado4"
   TextField "Campo de texto_8" at 233,557 size 155x18; Text 'Posición para Herramienta 1'
   GraphicView "Visor de gráficos_1" at 701,252 size 114x83; Picture "a_4"
   GraphicView "Visor de gráficos_2" at 972,251 size 114x83; Picture "b_2"
   GraphicView "Visor de gráficos_3" at 1022,197 size 114x83; Picture "c_1"
   GraphicView "Visor de gráficos_4" at 751,198 size 114x83; Picture "b_2"
   TextField "Campo de texto_22" at 857,426 size 41x18; Text 'Martillo'
      Visibility <- "MANU"
   TextField "Campo de texto_23" at 857,455 size 35x18; Text 'Matriz'
      Visibility <- "MANU"
   TextField "Campo de texto_24" at 1129,426 size 41x18; Text 'Martillo'
      Visibility <- "MANU"
   TextField "Campo de texto_25" at 1129,455 size 35x18; Text 'Matriz'
      Visibility <- "MANU"
   TextField "Campo de texto_3" at 504,662 size 51x18; Text 'Corner 1'
   TextField "Campo de texto_6" at 233,589 size 155x18; Text 'Posición para Herramienta 2'
   TextField "Campo de texto_7" at 812,557 size 155x18; Text 'Posición para Herramienta 1'
   TextField "Campo de texto_10" at 812,589 size 155x18; Text 'Posición para Herramienta 2'
   TextField "Campo de texto_11" at 731,661 size 51x18; Text 'Corner 2'
   TextField "Campo de texto_12" at 394,557 size 80x18; Text 'Ajuste con F1'
   TextField "Campo de texto_13" at 394,589 size 80x18; Text 'Ajuste con F2'
   TextField "Campo de texto_26" at 970,557 size 80x18; Text 'Ajuste con F3'
   TextField "Campo de texto_27" at 970,589 size 80x18; Text 'Ajuste con F4'

PopupScreen "Comandos Perfiladores" 1280x714
   Button "Botón_6" at 630,585 size 88x33; TextOff 'Avance'
      on Press: SetTag("DB_OP.RC1", 52); SetBit("DB_OP.OP_SELMANU1")
      Visibility <- "MANU"
      Appearance <- "DB_OP.RC1"
   Button "Botón_7" at 630,630 size 88x33; TextOff 'Retroceso'
      on Press: SetTag("DB_OP.RC1", 53); SetBit("DB_OP.OP_SELMANU1")
      Visibility <- "MANU"
      Appearance <- "DB_OP.RC1"
   Button "Botón_8" at 731,585 size 88x33; TextOff 'Hacia Consigna'
      on Press: SetTag("DB_OP.RC1", 51); SetBit("DB_OP.OP_SELMANU1")
      Visibility <- "MANU"
      Appearance <- "DB_OP.RC1"
   Button "Botón_11" at 731,630 size 88x33; TextOff 'Freno'
      on Press: SetTag("DB_OP.RC1", 54); SetBit("DB_OP.OP_SELMANU1")
      Visibility <- "MANU"
      Appearance <- "DB_OP.RC1"
   Button "Botón_1" at 889,270 size 88x33; TextOff 'Avance'
      on Press: SetTag("DB_OP.RC1", 55); SetBit("DB_OP.OP_SELMANU1")
      Visibility <- "MANU"
      Appearance <- "DB_OP.RC1"
   Button "Botón_2" at 889,307 size 88x33; TextOff 'Retroceso'
      on Press: SetTag("DB_OP.RC1", 56); SetBit("DB_OP.OP_SELMANU1")
      Visibility <- "MANU"
      Appearance <- "DB_OP.RC1"
   IOField "Champ E/S_1" at 943,573 size 77x29; FormatPattern 9999999
      ProcessValue <- "DB_OP.COD1_VAL"
   IOField "Champ E/S" at 947,636 size 70x29; FormatPattern 9.9999
      ProcessValue <- "DB_OP.COD1_COEF"
   IOField "Champ E/S_0" at 943,601 size 77x29; FormatPattern 9999999
      ProcessValue <- "DB_OP.COD1_CONS"
   IOField "Champ E/S_2" at 1114,575 size 69x29; FormatPattern 9999999
      ProcessValue <- "DB_OP.COD1_INIT"
   TextField "Champ de texte_2" at 861,578 size 82x18; Text 'Posición / Position Réelle'
   TextField "Champ de texte" at 844,607 size 99x18; Text 'Consigna / Position Consigne'
   TextField "Champ de texte_0" at 851,641 size 92x18; Text 'Coef corrección / Coeff correction'
   IOField "Champ E/S_4" at 1114,640 size 69x29; FormatPattern 9999999
      ProcessValue <- "DB_OP.COD1_TARGET"
   TextField "Champ de texte_5" at 1044,612 size 62x18; Text 'Cota Paro / Côte Arrêt'
   TextField "Champ de texte_6" at 1052,645 size 50x18; Text 'Ventana / Fenetre'
   IOField "Champ E/S_5" at 1114,607 size 69x29; FormatPattern 9999999
      ProcessValue <- "DB_OP.COD1_ARRET"
   Button "Button" at 1045,578 size 60x23; TextOff 'OFFSET'; Authorization "Nivel 1"
      on Press: SetBit("DB_OP.COD1_CMD")
      Appearance <- "DB_OP.COD2_CMD"
   GraphicIOField "Campo ES gráfico_4" at 236,203 size 456x232; PictureList "Grupo 2 - Perfilador"
      ProcessValue <- "Alarma_Perfiladores"
   Polygon "Polígono_3" at 265,240 size 389x46
      Visibility <- "Perfiladores\Perfilador.PresenciaPieza"
   Rectangle "Rectángulo_2" at 874,227 size 118x128
      Visibility <- "MANU"
   Rectangle "Rectángulo_3" at 874,227 size 118x29
      Visibility <- "MANU"
   TextField "Campo de texto_1" at 900,231 size 66x18; Text 'Perfiladores'
      Visibility <- "MANU"
   Circle "Cercle_11" at 450,253 size 12x12
      Appearance <- "27S4"
   Circle "Cercle_12" at 413,405 size 12x12
      Appearance <- "29S7"
   Circle "Cercle_13" at 411,387 size 12x12
      Appearance <- "29S7"
   Circle "Cercle_14" at 515,384 size 12x12
      Appearance <- "23S4"
   Polygon "Polígono_1" at 248,269 size 17x19
      Appearance <- "36S70"
   TextField "Campo de texto_3" at 246,143 size 112x18; Text 'Sensores de Atasco'
   TextField "Campo de texto_4" at 613,454 size 141x18; Text '23S4 - Presión de Frenos'
   TextField "Campo de texto_5" at 414,107 size 101x18; Text 'Motor Perfilador 4'
   TextField "Campo de texto_6" at 684,429 size 101x18; Text 'Motor Perfilador 3'
   TextField "Campo de texto_7" at 159,441 size 101x18; Text 'Motor Perfilador 1'
   TextField "Campo de texto_8" at 147,165 size 101x18; Text 'Motor Perfilador 2'
   TextField "Campo de texto_9" at 140,188 size 64x46; Text '36S70 Barrera de Atascos'
   TextField "Campo de texto_10" at 557,500 size 197x18; Text 'M07 - Motor Ajuste de Profundidad'
   TextField "Campo de texto_11" at 202,476 size 119x18; Text '29S7 - Fin de Carrera'
   TextField "Campo de texto_13" at 320,502 size 53x18; Text 'Encóder'
   TextField "Campo de texto_14" at 118,363 size 81x46; Text '27S3 - Chapa en Entrada Perfilador'
   Circle "Cercle_2" at 236,274 size 12x12
      Appearance <- "27S3"
   Polyline "Línea poligonal_11" at 263,255 size 397x22
      Appearance <- "36S70"
   Polygon "Polígono_2" at 655,246 size 17x19
      Appearance <- "36S70"
   Rectangle "Rectángulo_6" at 613,555 size 222x128
      Visibility <- "MANU"
   Rectangle "Rectángulo_7" at 834,539 size 374x144
      Visibility <- "MANU"
   Rectangle "Rectángulo_8" at 613,539 size 595x29
      Visibility <- "MANU"
   TextField "Campo de texto_12" at 674,543 size 108x18; Text 'Ajuste Profundidad'
      Visibility <- "MANU"

PopupScreen "Comandos Cinta" 1280x714
   Button "Botón_6" at 630,585 size 88x33; TextOff 'Avance'
      on Press: SetTag("DB_OP.RC1", 52); SetBit("DB_OP.OP_SELMANU1")
      Visibility <- "MANU"
      Appearance <- "DB_OP.RC1"
   Button "Botón_7" at 630,630 size 88x33; TextOff 'Retroceso'
      on Press: SetTag("DB_OP.RC1", 53); SetBit("DB_OP.OP_SELMANU1")
      Visibility <- "MANU"
      Appearance <- "DB_OP.RC1"
   Button "Botón_8" at 731,585 size 88x33; TextOff 'Hacia Consigna'
      on Press: SetTag("DB_OP.RC1", 51); SetBit("DB_OP.OP_SELMANU1")
      Visibility <- "MANU"
      Appearance <- "DB_OP.RC1"
   Button "Botón_11" at 731,630 size 88x33; TextOff 'Freno'
      on Press: SetTag("DB_OP.RC1", 54); SetBit("DB_OP.OP_SELMANU1")
      Visibility <- "MANU"
      Appearance <- "DB_OP.RC1"
   Button "Botón_4" at 462,582 size 88x33; TextOff 'Avance'
      on Press: SetTag("DB_OP.RC2", 91); SetBit("DB_OP.OP_SELMANU2")
      Visibility <- "MANU"
      Appearance <- "DB_OP.RC2"
   Button "Botón_5" at 462,619 size 88x33; TextOff 'Retroceso'
      on Press: SetTag("DB_OP.RC2", 92); SetBit("DB_OP.OP_SELMANU2")
      Visibility <- "MANU"
      Appearance <- "DB_OP.RC2"
   IOField "Champ E/S_1" at 943,573 size 77x29; FormatPattern 9999999
      ProcessValue <- "DB_OP.COD2_VAL"
   IOField "Champ E/S" at 947,636 size 70x29; FormatPattern 9.9999
      ProcessValue <- "DB_OP.COD2_COEF"
   IOField "Champ E/S_0" at 943,601 size 77x29; FormatPattern 9999999
      ProcessValue <- "DB_OP.COD2_CONS"
   IOField "Champ E/S_2" at 1114,575 size 69x29; FormatPattern 9999999
      ProcessValue <- "DB_OP.COD2_INIT"
   TextField "Champ de texte_2" at 861,578 size 82x18; Text 'Posición / Position Réelle'
   TextField "Champ de texte" at 844,607 size 99x18; Text 'Consigna / Position Consigne'
   TextField "Champ de texte_0" at 851,641 size 92x18; Text 'Coef corrección / Coeff correction'
   IOField "Champ E/S_4" at 1114,640 size 69x29; FormatPattern 9999999
      ProcessValue <- "DB_OP.COD2_TARGET"
   TextField "Champ de texte_5" at 1044,612 size 62x18; Text 'Cota Paro / Côte Arrêt'
   TextField "Champ de texte_6" at 1052,645 size 50x18; Text 'Ventana / Fenetre'
   IOField "Champ E/S_5" at 1114,607 size 69x29; FormatPattern 9999999
      ProcessValue <- "DB_OP.COD2_ARRET"
   Button "Button" at 1045,578 size 60x23; TextOff 'OFFSET'; Authorization "Nivel 1"
      on Press: SetBit("DB_OP.COD2_CMD")
      Appearance <- "DB_OP.COD2_CMD"
   GraphicIOField "Campo ES gráfico_1" at 290,222 size 647x180; PictureList "Grupo 2 - Cinta"
      ProcessValue <- "Alarma_Cinta"
   Rectangle "Rectángulo_1" at 613,555 size 222x128
      Visibility <- "MANU"
   Rectangle "Rectángulo_2" at 448,539 size 118x128
      Visibility <- "MANU"
   Rectangle "Rectángulo_3" at 448,539 size 118x29
      Visibility <- "MANU"
   TextField "Campo de texto_1" at 474,543 size 31x18; Text 'Cinta'
      Visibility <- "MANU"
   Rectangle "Rectángulo_6" at 834,539 size 374x144
      Visibility <- "MANU"
   Rectangle "Rectángulo_7" at 613,539 size 595x29
      Visibility <- "MANU"
   TextField "Campo de texto_12" at 642,543 size 108x18; Text 'Ajuste Profundidad'
      Visibility <- "MANU"
   Circle "Cercle_1" at 325,248 size 12x12
      Appearance <- "27S4"
   Circle "Cercle_14" at 909,220 size 12x12
      Appearance <- "29S1"
   Circle "Cercle_15" at 909,234 size 12x12
      Appearance <- "29S2"
   Circle "Cercle_11" at 826,289 size 12x12
      Appearance <- "25S2"
   Circle "Cercle" at 911,284 size 12x12
      Appearance <- "29S3"
   TextField "Campo de texto_22" at 109,219 size 183x18; Text '27S4 - Chapa en Salida Perfilador'
   TextField "Campo de texto_23" at 624,433 size 179x18; Text 'M07 - Motor Ajuste Profundidad'
   TextField "Campo de texto_24" at 987,328 size 126x18; Text '25S2 - Bajar Velocidad'
   TextField "Campo de texto_25" at 512,385 size 223x18; Text '29S3 - Presencia de Chapa en Formador'
   TextField "Campo de texto_31" at 616,197 size 166x18; Text 'M08 - Motor Transporte Cinta'
   TextField "Campo de texto_32" at 667,130 size 145x18; Text '29S1 - Avance Bloqueado'
   TextField "Campo de texto_33" at 647,164 size 165x18; Text '29S2 - Avance Desbloqueado'
   Polygon "Polígono_4" at 351,252 size 385x62
      Visibility <- "Cinta\Cinta.PresenciaPieza"

